// TIA Portal project "Task 1 Faceplate" (V16)

(* hardware
DEVICE "S7-1200 station_1"  S7-1200 Station
   slot 0: "Rack_0"  S7-1200 Rack  Rack  V1.0
   slot 1: "PLC_1"  CPU 1215C DC/DC/DC  6ES7 215-1AG40-0XB0  V4.4
DEVICE "HMI_1"  TP700 Comfort
   slot 0: "HMI_1"  TP700 Comfort  6AV2 124-0GC01-0AX0  16.0.0.0
   slot 1: "HMI_RT_1"  TP700 Comfort  6AV2 124-0GC01-0AX0  16.0.0.0
   slot 5: "HMI_1.IE_CP_1"  PROFINET Interface  16.0.0.0
      slot 1: "PROFINET Interface_1"  PROFINET Interface
         slot 1: "Port_1"  Port
         slot 2: "Port_2"  Port
   slot 7: "HMI_1.MPI/DP_CP_1"  MPI/DP Interface  16.0.0.0
*)

// ===== PLC "PLC_1"  CPU 1215C DC/DC/DC =====

DATA_BLOCK "TASK2 FB"   // DB1
{ S7_Optimized_Access := 'TRUE' }
VERSION : 0.1
// stored: InstanceOfName TASK2
"TASK2"
BEGIN
END_DATA_BLOCK

DATA_BLOCK "TASK1 FB"   // DB2
{ S7_Optimized_Access := 'TRUE' }
VERSION : 0.1
// stored: InstanceOfName TASK1
"TASK1"
BEGIN
END_DATA_BLOCK

DATA_BLOCK "TASK1 DB"   // DB3
{ S7_Optimized_Access := 'TRUE' }
VERSION : 0.1
   VAR
      start : Bool;
      stop : Bool;
      heater : Bool;
   END_VAR
   VAR RETAIN
      temperature : Real;
   END_VAR
   VAR
      run : Bool;
      "max temp" : Real := 50.0;
      "min temp" : Real := 0.0;
      "reset temp" : Real := 0.0;
      reset : Bool;
   END_VAR
   VAR RETAIN
      "preset timer" : DInt := 1000;
   END_VAR
   VAR
      "max limit" : Bool;
      "min limit" : Bool;
      timer_1 : IEC_TIMER;
   END_VAR
BEGIN
END_DATA_BLOCK

DATA_BLOCK "TASK2 DB"   // DB4
{ S7_Optimized_Access := 'TRUE' }
VERSION : 0.1
   VAR
      START : Bool;
      STOP : Bool;
      RUN : Bool;
      FVV : Real := 0.0;
      DVV : Real := 0.0;
      "TIMER" : IEC_TIMER;
      "PRESET TIMER" : Real;
      "MULTIPLY BY X" : Real;
      "MAX LIQUID" : Real := 100.0;
      "MIN LIQUID" : Real := 0.0;
      "H LIQUID ALARM" : Real := 100.0;
      "L LIQUID ALARM" : Real := 20.0;
   END_VAR
BEGIN
END_DATA_BLOCK

FUNCTION_BLOCK "TASK1"   // FB1, LAD
{ S7_Optimized_Access := 'TRUE' }
VERSION : 0.1
   VAR_INPUT
      Start : Bool;
      Stop : Bool;
      reset : Bool;
      "Timer" : DInt;   // value in milliseconds
      "max temperature" : Real;   // max temperature you want in the tank
      "min temperature" : Real;   // min temperature you want in the tank
      "reset temp" : Real;   // to reset the temperature
      "any value" : Real;
      manual : Bool;
   END_VAR
   VAR_OUTPUT
      Output_1 : Bool;
   END_VAR
   VAR_IN_OUT
      Run : Bool;   // process is working
      Heater : Bool;
      "max limit" : Bool;
      "min limit" : Bool;
      Temperature : Real;
      IEC_Timer_0_Instance : TON_TIME;
   END_VAR
   VAR
      Ton : Bool;
      Toff : Bool;   // reset the timer
   END_VAR
BEGIN

REGION Network 1: control operarion
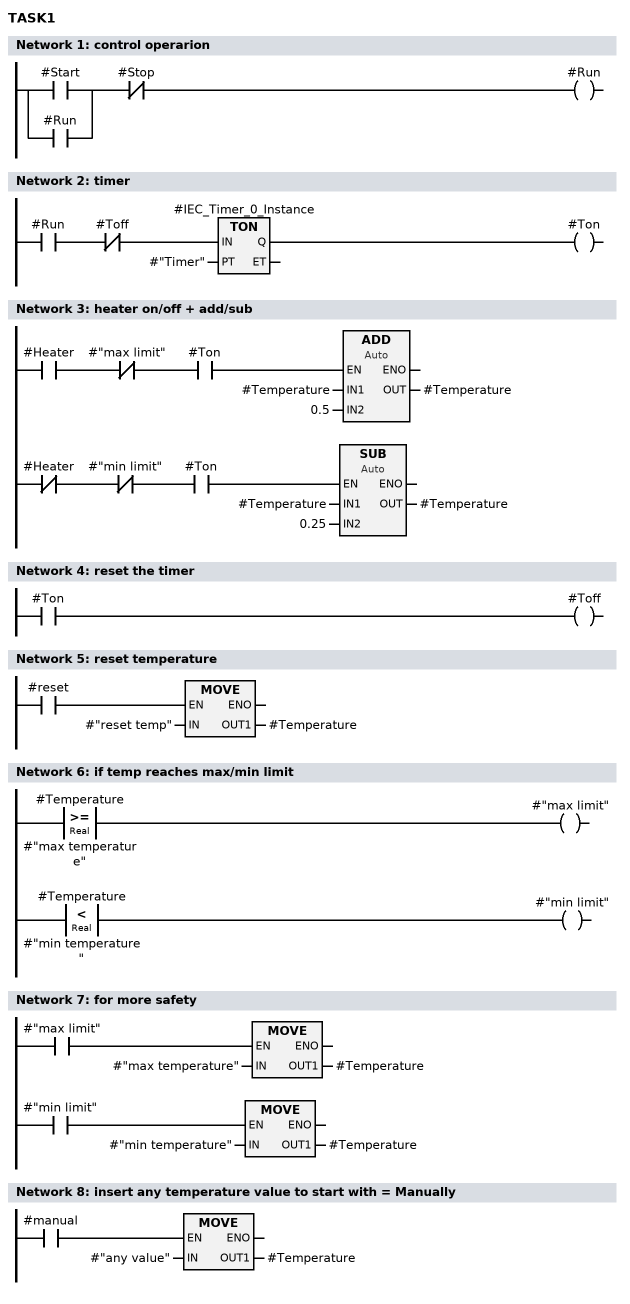
   RUNG wire#powerrail
      Contact( #Start )
      wire#w1
      I_Contact( #Stop )
      Coil( #Run )
   END_RUNG
   RUNG wire#powerrail
      Contact( #Run )
   END_RUNG wire#w1
   // the same network as SCL:
   #Run := (#Start OR #Run) AND NOT #Stop;
END_REGION

REGION Network 2: timer
   #IEC_Timer_0_Instance(IN := #Run AND NOT #Toff, PT := #"Timer");   // TON
   #Ton := #IEC_Timer_0_Instance.Q;
END_REGION

REGION Network 3: heater on/off + add/sub
   RUNG wire#powerrail
      Contact( #Heater )
      I_Contact( #"max limit" )
      Contact( #Ton )
      Add(in1 := #Temperature, in2 := 0.5, out => #Temperature)
   END_RUNG
   RUNG wire#powerrail
      I_Contact( #Heater )
      I_Contact( #"min limit" )
      Contact( #Ton )
      Sub(in1 := #Temperature, in2 := 0.25, out => #Temperature)
   END_RUNG
   // the same network as SCL:
   IF #Heater AND NOT #"max limit" AND #Ton THEN #Temperature := #Temperature + 0.5; END_IF;
   IF NOT #Heater AND NOT #"min limit" AND #Ton THEN #Temperature := #Temperature - 0.25; END_IF;
END_REGION

REGION Network 4: reset the timer
   RUNG wire#powerrail
      Contact( #Ton )
      Coil( #Toff )
   END_RUNG
   // the same network as SCL:
   #Toff := #Ton;
END_REGION

REGION Network 5: reset temperature
   RUNG wire#powerrail
      Contact( #reset )
      Move(in := #"reset temp", out1 => #Temperature)
   END_RUNG
   // the same network as SCL:
   IF #reset THEN #Temperature := #"reset temp"; END_IF;
END_REGION

REGION Network 6: if temp reaches max/min limit
   RUNG wire#powerrail
      { S7_Templates := "SrcType := Real" } GE_Contact(in1 := #Temperature, in2 := #"max temperature")
      Coil( #"max limit" )
   END_RUNG
   RUNG wire#powerrail
      { S7_Templates := "SrcType := Real" } LT_Contact(in1 := #Temperature, in2 := #"min temperature")
      Coil( #"min limit" )
   END_RUNG
   // the same network as SCL:
   #"max limit" := #Temperature >= #"max temperature";
   #"min limit" := #Temperature < #"min temperature";
END_REGION

REGION Network 7: for more safety
   RUNG wire#powerrail
      Contact( #"max limit" )
      Move(in := #"max temperature", out1 => #Temperature)
   END_RUNG
   RUNG wire#powerrail
      Contact( #"min limit" )
      Move(in := #"min temperature", out1 => #Temperature)
   END_RUNG
   // the same network as SCL:
   IF #"max limit" THEN #Temperature := #"max temperature"; END_IF;
   IF #"min limit" THEN #Temperature := #"min temperature"; END_IF;
END_REGION

REGION Network 8: insert any temperature value to start with = Manually
   RUNG wire#powerrail
      Contact( #manual )
      Move(in := #"any value", out1 => #Temperature)
   END_RUNG
   // the same network as SCL:
   IF #manual THEN #Temperature := #"any value"; END_IF;
END_REGION
END_FUNCTION_BLOCK

FUNCTION_BLOCK "TASK2"   // FB2, LAD
{ S7_Optimized_Access := 'TRUE' }
VERSION : 0.1
   VAR_INPUT
      start : Bool;
      stop : Bool;
      "fill valve voltage" : Real;   // analog input from 0-10v
      "drain valve voltage" : Real;   // analog input from 0-10v
      "multiply by x" : Real;   // your max value
      "TIMER" : DInt;   // TIME IN MILLISECONDS FOR CHANGE
      "HIGH LIQUID ALARM" : Real;
      "LOW LIQUID ALARM" : Real;
   END_VAR
   VAR_OUTPUT
      "REAL FVV" : Real;   // real fill valve voltage
      "REAL DVV" : Real;   // real drain valve voltage
      "HIGH LEVEL ALARM" : Bool;
      "LOW LEVEL ALARM" : Bool;
   END_VAR
   VAR_IN_OUT
      run : Bool;
      Rate : Real;   // FLOW OF LIQUID PER TIME
      "REAL FVV - REAL DVV" : Real;
      IEC_Timer_0_Instance : TON_TIME;
      "MAX LEVEL" : Bool;
      "MIN LEVEL" : Bool;
      LEVEL : Real;   // LEVEL OF THE LIQUID
      "MAX LIQUID" : Real;   // MAX LEVEL LIQUID ACCEPTED
      "MIN LIQUID" : Real;   // MIN LEVEL LIQUID ACCEPTED
   END_VAR
   VAR
      "division by 10" : Real := 10.0;
      "FVV after division" : Real;
      "DVV after division" : Real;
      TON : Bool;
      TOFF : Bool;
   END_VAR
BEGIN

REGION Network 1: control process
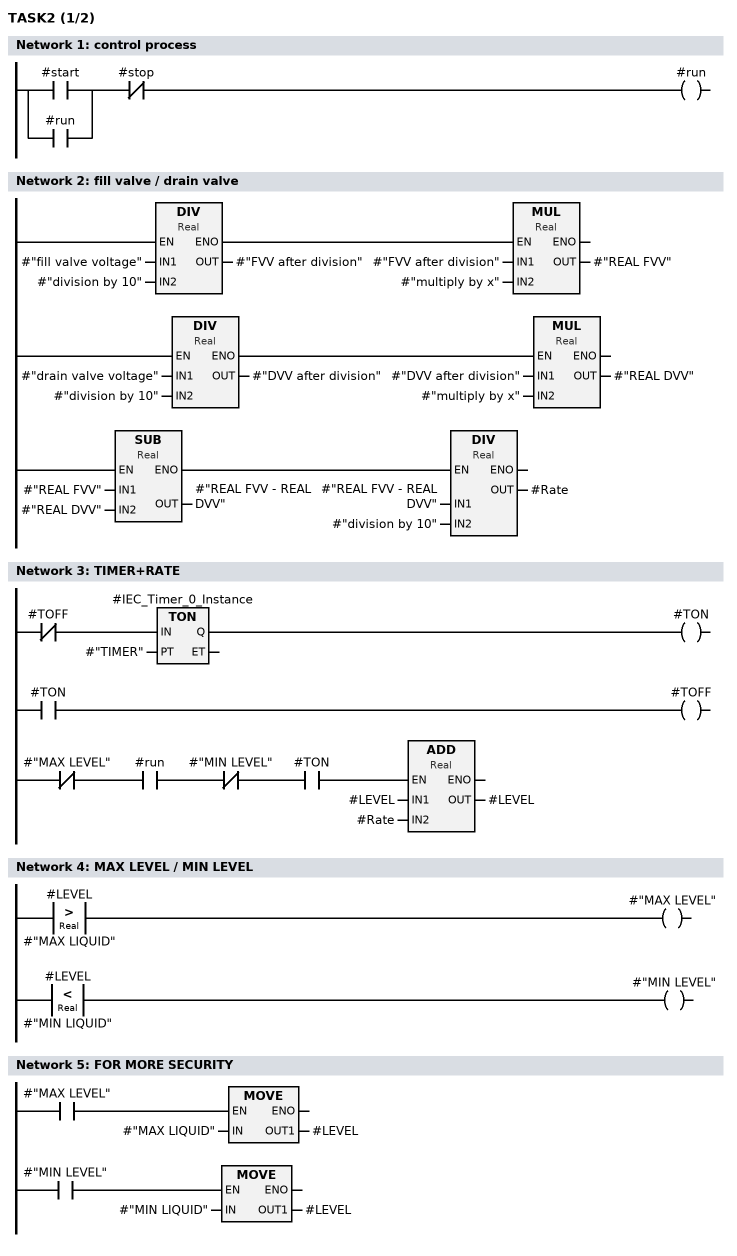
   RUNG wire#powerrail
      Contact( #start )
      wire#w1
      I_Contact( #stop )
      Coil( #run )
   END_RUNG
   RUNG wire#powerrail
      Contact( #run )
   END_RUNG wire#w1
   // the same network as SCL:
   #run := (#start OR #run) AND NOT #stop;
END_REGION

REGION Network 2: fill valve / drain valve
   RUNG wire#powerrail
      { S7_Templates := "SrcType := Real" } Div(in1 := #"fill valve voltage", in2 := #"division by 10", out => #"FVV after division")
      { S7_Templates := "SrcType := Real" } Mul(in1 := #"FVV after division", in2 := #"multiply by x", out => #"REAL FVV")
   END_RUNG
   RUNG wire#powerrail
      { S7_Templates := "SrcType := Real" } Div(in1 := #"drain valve voltage", in2 := #"division by 10", out => #"DVV after division")
      { S7_Templates := "SrcType := Real" } Mul(in1 := #"DVV after division", in2 := #"multiply by x", out => #"REAL DVV")
   END_RUNG
   RUNG wire#powerrail
      { S7_Templates := "SrcType := Real" } Sub(in1 := #"REAL FVV", in2 := #"REAL DVV", out => #"REAL FVV - REAL DVV")
      { S7_Templates := "SrcType := Real" } Div(in1 := #"REAL FVV - REAL DVV", in2 := #"division by 10", out => #Rate)
   END_RUNG
   // the same network as SCL:
   #"FVV after division" := #"fill valve voltage" / #"division by 10";
   #"REAL FVV" := #"FVV after division" * #"multiply by x";
   #"DVV after division" := #"drain valve voltage" / #"division by 10";
   #"REAL DVV" := #"DVV after division" * #"multiply by x";
   #"REAL FVV - REAL DVV" := #"REAL FVV" - #"REAL DVV";
   #Rate := #"REAL FVV - REAL DVV" / #"division by 10";
END_REGION

REGION Network 3: TIMER+RATE
   #IEC_Timer_0_Instance(IN := NOT #TOFF, PT := #"TIMER");   // TON
   #TON := #IEC_Timer_0_Instance.Q;
   #TOFF := #TON;
   IF NOT #"MAX LEVEL" AND #run AND NOT #"MIN LEVEL" AND #TON THEN #LEVEL := #LEVEL + #Rate; END_IF;
END_REGION

REGION Network 4: MAX LEVEL / MIN LEVEL
   RUNG wire#powerrail
      { S7_Templates := "SrcType := Real" } GT_Contact(in1 := #LEVEL, in2 := #"MAX LIQUID")
      Coil( #"MAX LEVEL" )
   END_RUNG
   RUNG wire#powerrail
      { S7_Templates := "SrcType := Real" } LT_Contact(in1 := #LEVEL, in2 := #"MIN LIQUID")
      Coil( #"MIN LEVEL" )
   END_RUNG
   // the same network as SCL:
   #"MAX LEVEL" := #LEVEL > #"MAX LIQUID";
   #"MIN LEVEL" := #LEVEL < #"MIN LIQUID";
END_REGION

REGION Network 5: FOR MORE SECURITY
   RUNG wire#powerrail
      Contact( #"MAX LEVEL" )
      Move(in := #"MAX LIQUID", out1 => #LEVEL)
   END_RUNG
   RUNG wire#powerrail
      Contact( #"MIN LEVEL" )
      Move(in := #"MIN LIQUID", out1 => #LEVEL)
   END_RUNG
   // the same network as SCL:
   IF #"MAX LEVEL" THEN #LEVEL := #"MAX LIQUID"; END_IF;
   IF #"MIN LEVEL" THEN #LEVEL := #"MIN LIQUID"; END_IF;
END_REGION

REGION Network 6: HIGH LEVEL ALARM / LOW LEVEL ALARM
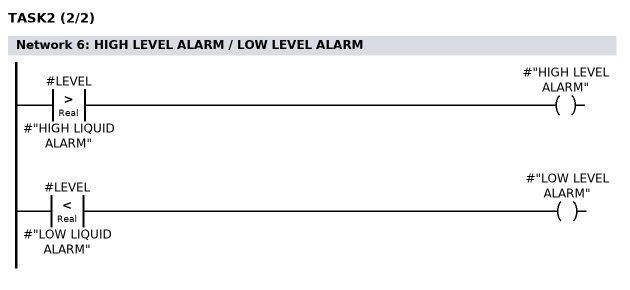
   RUNG wire#powerrail
      { S7_Templates := "SrcType := Real" } GT_Contact(in1 := #LEVEL, in2 := #"HIGH LIQUID ALARM")
      Coil( #"HIGH LEVEL ALARM" )
   END_RUNG
   RUNG wire#powerrail
      { S7_Templates := "SrcType := Real" } LT_Contact(in1 := #LEVEL, in2 := #"LOW LIQUID ALARM")
      Coil( #"LOW LEVEL ALARM" )
   END_RUNG
   // the same network as SCL:
   #"HIGH LEVEL ALARM" := #LEVEL > #"HIGH LIQUID ALARM";
   #"LOW LEVEL ALARM" := #LEVEL < #"LOW LIQUID ALARM";
END_REGION
END_FUNCTION_BLOCK

ORGANIZATION_BLOCK "Main"   // OB1, LAD, ProgramCycle
TITLE = "Main Program Sweep (Cycle)"
{ S7_Optimized_Access := 'TRUE' }
VERSION : 0.1
   VAR_INPUT
      Initial_Call : Bool;   // Initial call of this OB
      Remanence : Bool;   // =True, if remanent data are available
   END_VAR
BEGIN

REGION Network 1
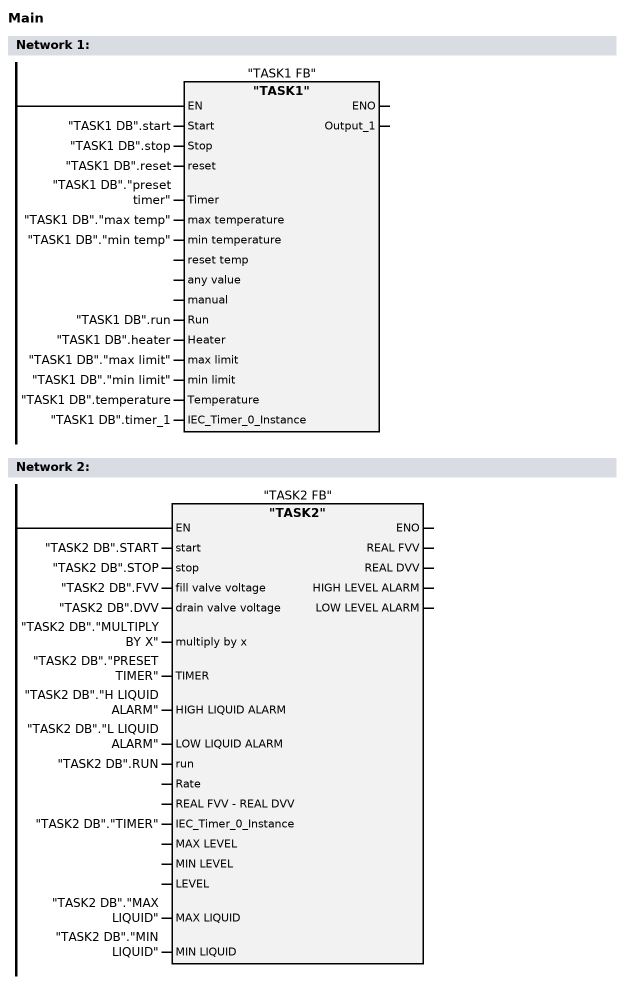
   RUNG wire#powerrail
      "TASK1 FB"(Start := "TASK1 DB".start, Stop := "TASK1 DB".stop, reset := "TASK1 DB".reset, "Timer" := "TASK1 DB"."preset timer", "max temperature" := "TASK1 DB"."max temp", "min temperature" := "TASK1 DB"."min temp", "reset temp" :=, "any value" :=, manual :=, Run := "TASK1 DB".run, Heater := "TASK1 DB".heater, "max limit" := "TASK1 DB"."max limit", "min limit" := "TASK1 DB"."min limit", Temperature := "TASK1 DB".temperature, IEC_Timer_0_Instance := "TASK1 DB".timer_1, Output_1 =>)
   END_RUNG
   // the same network as SCL:
   "TASK1 FB"(Start := "TASK1 DB".start,   // "TASK1"
              Stop := "TASK1 DB".stop,
              reset := "TASK1 DB".reset,
              "Timer" := "TASK1 DB"."preset timer",
              "max temperature" := "TASK1 DB"."max temp",
              "min temperature" := "TASK1 DB"."min temp",
              Run := "TASK1 DB".run,
              Heater := "TASK1 DB".heater,
              "max limit" := "TASK1 DB"."max limit",
              "min limit" := "TASK1 DB"."min limit",
              Temperature := "TASK1 DB".temperature,
              IEC_Timer_0_Instance := "TASK1 DB".timer_1);
END_REGION

REGION Network 2
   RUNG wire#powerrail
      "TASK2 FB"(start := "TASK2 DB".START, stop := "TASK2 DB".STOP, "fill valve voltage" := "TASK2 DB".FVV, "drain valve voltage" := "TASK2 DB".DVV, "multiply by x" := "TASK2 DB"."MULTIPLY BY X", "TIMER" := "TASK2 DB"."PRESET TIMER", "HIGH LIQUID ALARM" := "TASK2 DB"."H LIQUID ALARM", "LOW LIQUID ALARM" := "TASK2 DB"."L LIQUID ALARM", run := "TASK2 DB".RUN, Rate :=, "REAL FVV - REAL DVV" :=, IEC_Timer_0_Instance := "TASK2 DB"."TIMER", "MAX LEVEL" :=, "MIN LEVEL" :=, LEVEL :=, "MAX LIQUID" := "TASK2 DB"."MAX LIQUID", "MIN LIQUID" := "TASK2 DB"."MIN LIQUID", "REAL FVV" =>, "REAL DVV" =>, "HIGH LEVEL ALARM" =>, "LOW LEVEL ALARM" =>)
   END_RUNG
   // the same network as SCL:
   "TASK2 FB"(start := "TASK2 DB".START,   // "TASK2"
              stop := "TASK2 DB".STOP,
              "fill valve voltage" := "TASK2 DB".FVV,
              "drain valve voltage" := "TASK2 DB".DVV,
              "multiply by x" := "TASK2 DB"."MULTIPLY BY X",
              "TIMER" := "TASK2 DB"."PRESET TIMER",
              "HIGH LIQUID ALARM" := "TASK2 DB"."H LIQUID ALARM",
              "LOW LIQUID ALARM" := "TASK2 DB"."L LIQUID ALARM",
              run := "TASK2 DB".RUN,
              IEC_Timer_0_Instance := "TASK2 DB"."TIMER",
              "MAX LIQUID" := "TASK2 DB"."MAX LIQUID",
              "MIN LIQUID" := "TASK2 DB"."MIN LIQUID");
END_REGION
END_ORGANIZATION_BLOCK

// ===== library: MasterCopy "TASK1 DB" =====

DATA_BLOCK "TASK1 DB"   // DB3
{ S7_Optimized_Access := 'TRUE' }
VERSION : 0.1
   VAR
      start : Bool;
      stop : Bool;
      heater : Bool;
   END_VAR
   VAR RETAIN
      temperature : Real;
   END_VAR
   VAR
      run : Bool;
      "max temp" : Real := 50.0;
      "min temp" : Real := 0.0;
      "reset temp" : Real := 0.0;
      reset : Bool;
   END_VAR
   VAR RETAIN
      "preset timer" : DInt := 1000;
   END_VAR
   VAR
      "max limit" : Bool;
      "min limit" : Bool;
      timer_1 : IEC_TIMER;
   END_VAR
BEGIN
END_DATA_BLOCK

// ===== library: MasterCopy "TASK2 DB" =====

DATA_BLOCK "TASK2 DB"   // DB4
{ S7_Optimized_Access := 'TRUE' }
VERSION : 0.1
   VAR
      START : Bool;
      STOP : Bool;
      RUN : Bool;
      FVV : Real := 0.0;
      DVV : Real := 0.0;
      "TIMER" : IEC_TIMER;
      "PRESET TIMER" : Real;
      "MULTIPLY BY X" : Real;
      "MAX LIQUID" : Real := 100.0;
      "MIN LIQUID" : Real := 0.0;
      "H LIQUID ALARM" : Real := 100.0;
      "L LIQUID ALARM" : Real := 20.0;
   END_VAR
BEGIN
END_DATA_BLOCK

(* ===== HMI "HMI_RT_1" =====
system functions are stored by id; their names below are inferred from use
connection "HMI_Connection_1": ETHERNET, S7_1200_OMS

HMI tags "Default tag table"
   "Tag_ScreenNumber" : UInt, internal
   "Data_block_1_temperature" : Real = PLC "TASK1 DB".temperature, 1 s
   "Data_block_1_start" : Bool = PLC "TASK1 DB".start, 1 s
   "Data_block_1_heater" : Bool = PLC "TASK1 DB".heater, 1 s
   "TASK1 DB_stop" : Bool = PLC "TASK1 DB".stop, 1 s
   "TASK1 DB_reset" : Bool = PLC "TASK1 DB".reset, 1 s

Template "Template_1" 800x480
   Button "Exit" at 714,429 size 71x50; TextOff 'Exit'; PictureOff "ExitRuntime_KTP700_Basic_PN_TR"; PictureOn "ExitRuntime_KTP700_Basic_PN_TR"
      on Release: StopRuntime(0)
   Button "Template_Button" at 614,429 size 71x50; TextOff 'Text'
   Button "Template_Button_1" at 514,429 size 71x50; TextOff 'Text'
   Button "Template_Button_2" at 414,429 size 71x50; TextOff 'Text'
   Button "Template_Button_3" at 314,429 size 71x50; TextOff 'Text'
   Button "Template_Button_4" at 214,429 size 71x50; TextOff 'Text'
   Button "Template_Button_5" at 114,429 size 71x50; TextOff 'Text'
   Button "Start screen" at 14,429 size 71x50; TextOff 'Start screen'; PictureOff "NavigateHome_KTP700_Basic_PN_TR"; PictureOn "NavigateHome_KTP700_Basic_PN_TR"
      on Release: ActivateScreen("Root screen", 0)
   SymbolicIOField "Symbolic_IO_Field_Screen" at 93,9 size 600x33; TextOff '0'; TextOn '1'; TextList "TextList_ScreenNames"
      ProcessValue <- "Tag_ScreenNumber"
      on Change: ActivateScreenByNumber("Tag_ScreenNumber", 0)
   DateTimeField "HmiScreenItemData" at 695,25 size 105x25
   DateTimeField "HmiScreenItemData_1" at 695,0 size 105x25
   GraphicView "Logo" at 0,0 size 91x51; Picture "Logo of HMI_1"

screen "Root screen" 800x480, template "Template_1"
   on GenerateScreen: SetTag("Tag_ScreenNumber", 1)
   TextField "HmiScreenItemData" at 86,12 size 640x25; Text 'Welcome to HMI_1 (KTP700 Basic+ PN)!'
   ScreenModuleView "Faceplate_3_1" at 50,59 size 202x216; Guid_{11997190-8919} 'temp1'; ScreenModuleType ""; Guid_{11997190-9122} 'Temperature'
      Guid_{11997190-7705} <- "Data_block_1_heater"
      Guid_{11997190-7699} <- "Data_block_1_start"
      Guid_{11997190-7703} <- "TASK1 DB_stop"
      Guid_{11997190-7872} <- "Data_block_1_temperature"
      Guid_{11997190-7707} <- "TASK1 DB_reset"
   ScreenModuleView "Faceplate_3_2" at 297,56 size 202x216; ScreenModuleType ""
      Guid_{11997190-7705} <- "Data_block_1_heater"
*)

(* ===== HMI "HMI_RT_1" =====

ScreenModuleEditorView "Faceplate_3" 640x480
   Button "Button_2" at 14,148 size 96x32; TextOff 'Start'
   Button "Button_3" at 115,148 size 96x32; TextOff 'Stop'
   IOField "I/O field_1" at 31,56 size 165x32; FormatPattern s999.99
   Button "Button_4" at 53,17 size 116x32; TextOff 'Temperature'
   Switch "Switch_1" at 51,102 size 114x32; TextOn 'Heater ON'; CaptionText 'Switch'; TextOff 'Heater OFF'
   Button "Button_1" at 59,192 size 96x32; TextOff 'Reset'
*)

(* ===== HMI "HMI_RT_1" =====

ScreenModuleEditorView "Faceplate_3" 640x480
   Button "Button_2" at 14,148 size 96x32; TextOff 'Start'
   Button "Button_3" at 115,148 size 96x32; TextOff 'Stop'
   IOField "I/O field_1" at 31,56 size 165x32; FormatPattern s999.99
   Button "Button_4" at 53,17 size 116x32; TextOff 'Temperature'
   Switch "Switch_1" at 51,102 size 114x32; TextOn 'Heater ON'; CaptionText 'Switch'; TextOff 'Heater OFF'
   Button "Button_1" at 59,192 size 96x32; TextOff 'Reset'
*)

(* ===== HMI "HMI_RT_1" =====

ScreenModuleEditorView "Faceplate_3" 640x480
   Button "Button_2" at 14,148 size 96x32; TextOff 'Start'
   Button "Button_3" at 115,148 size 96x32; TextOff 'Stop'
   IOField "I/O field_1" at 31,56 size 165x32; FormatPattern s999.99
   Button "Button_4" at 53,17 size 116x32; TextOff 'Temperature'
   Switch "Switch_1" at 51,102 size 114x32; TextOn 'Heater ON'; CaptionText 'Switch'; TextOff 'Heater OFF'
   Button "Button_1" at 59,192 size 96x32; TextOff 'Reset'
*)

(* ===== HMI "HMI_RT_1" =====
system functions are stored by id; their names below are inferred from use

ScreenModuleEditorView "Faceplate_3" 640x480
   Button "Button_2" at 14,148 size 96x32; TextOff 'Start'
      on Press: SetBit("Start")
      on Release: ResetBit("Start")
   Button "Button_3" at 115,148 size 96x32; TextOff 'Stop'
      ProcessValue <- "stop"
      on Press: SetBit("stop")
      on Release: ResetBit("stop")
   IOField "I/O field_1" at 31,56 size 165x32; FormatPattern s99999
      ProcessValue <- "Temperature"
   Button "Button_4" at 44,17 size 130x32; TextOff 'Temperature'
   Switch "Switch_1" at 51,102 size 114x32; TextOn 'Heater ON'; CaptionText 'Switch'; TextOff 'Heater OFF'
      on SwitchOn: SetBit("Heater")
      on SwitchOff: ResetBit("Heater")
   Button "Button_1" at 59,192 size 96x32; TextOff 'Reset'
*)

(* ===== HMI "HMI_RT_1" =====
system functions are stored by id; their names below are inferred from use

ScreenModuleEditorView "Faceplate_3" 640x480
   Button "Button_2" at 14,148 size 96x32; TextOff 'Start'
      on Release: ResetBit("Start")
      on Press: SetBit("Start")
   Button "Button_3" at 115,148 size 96x32; TextOff 'Stop'
      on Release: ResetBit("stop")
      on Press: SetBit("stop")
      ProcessValue <- "stop"
   IOField "I/O field_1" at 31,56 size 165x32; FormatPattern s99999
      ProcessValue <- "Temperature"
   Button "Button_4" at 44,17 size 130x32; TextOff 'Temperature'
   Switch "Switch_1" at 51,102 size 114x32; TextOn 'Heater ON'; CaptionText 'Switch'; TextOff 'Heater OFF'
      on SwitchOff: ResetBit("Heater")
      on SwitchOn: SetBit("Heater")
   Button "Button_1" at 59,192 size 96x32; TextOff 'Reset'
*)

(* ===== HMI "HMI_RT_1" =====
system functions are stored by id; their names below are inferred from use

ScreenModuleEditorView "Faceplate_3" 640x480
   Button "Button_2" at 14,148 size 96x32; TextOff 'Start'
      on Release: ResetBit("Start")
      on Press: SetBit("Start")
      ProcessValue <- "Start"
   Button "Button_3" at 115,148 size 96x32; TextOff 'Stop'
      on Release: ResetBit("stop")
      on Press: SetBit("stop")
      ProcessValue <- "stop"
   IOField "I/O field_1" at 31,56 size 165x32; FormatPattern s99999
      ProcessValue <- "Temperature"
   Button "Button_4" at 44,17 size 130x32; TextOff 'Temperature'
   Switch "Switch_1" at 51,102 size 114x32; TextOn 'Heater ON'; CaptionText 'Switch'; TextOff 'Heater OFF'
      on SwitchOn: SetBit("Heater")
      on SwitchOff: ResetBit("Heater")
      ProcessValue <- "Heater"
   Button "Button_1" at 59,192 size 96x32; TextOff 'Reset'
      ProcessValue <- "reset"
*)

(* ===== HMI "HMI_RT_1" =====
system functions are stored by id; their names below are inferred from use

ScreenModuleEditorView "Faceplate_3" 640x480
   Button "Button_2" at 14,148 size 96x32; TextOff 'Start'
      on Release: ResetBit("Start")
      on Press: SetBit("Start")
      ProcessValue <- "Start"
   Button "Button_3" at 115,148 size 96x32; TextOff 'Stop'
      on Release: ResetBit("stop")
      on Press: SetBit("stop")
      ProcessValue <- "stop"
   IOField "I/O field_1" at 31,56 size 165x32; FormatPattern s999.99
      ProcessValue <- "Temperature"
   Button "Button_4" at 44,17 size 130x32; TextOff 'Temperature'
   Switch "Switch_1" at 51,102 size 114x32; TextOn 'Heater ON'; CaptionText 'Switch'; TextOff 'Heater OFF'
      on SwitchOff: ResetBit("Heater")
      on SwitchOn: SetBit("Heater")
      ProcessValue <- "Heater"
   Button "Button_1" at 59,192 size 96x32; TextOff 'Reset'
      ProcessValue <- "reset"
*)

(* ===== HMI "HMI_RT_1" =====
system functions are stored by id; their names below are inferred from use

ScreenModuleEditorView "Faceplate_3" 640x480
   Button "Button_2" at 14,148 size 96x32; TextOff 'Start'
      on Release: ResetBit("Start")
      on Press: SetBit("Start")
      ProcessValue <- "Start"
   Button "Button_3" at 115,148 size 96x32; TextOff 'Stop'
      on Release: ResetBit("stop")
      on Press: SetBit("stop")
      ProcessValue <- "stop"
   IOField "I/O field_1" at 31,56 size 165x32; FormatPattern s999.99
      ProcessValue <- "Temperature"
   Button "Button_4" at 44,17 size 130x32; TextOff 'Temperature'
   Switch "Switch_1" at 51,102 size 114x32; TextOn 'Heater ON'; CaptionText 'Switch'; TextOff 'Heater OFF'
      on SwitchOff: ResetBit("Heater")
      on SwitchOn: SetBit("Heater")
      ProcessValue <- "Heater"
   Button "Button_1" at 59,192 size 96x32; TextOff 'Reset'
      ProcessValue <- "reset"
      on Press: SetBit("reset")
      on Release: ResetBit("reset")
*)

(* ===== HMI "HMI_RT_1" =====
system functions are stored by id; their names below are inferred from use

ScreenModuleEditorView "Faceplate_3" 640x480
   Button "Button_2" at 14,148 size 96x32; TextOff 'Start'
      on Release: ResetBit("Start")
      on Press: SetBit("Start")
      ProcessValue <- "Start"
   Button "Button_3" at 115,148 size 96x32; TextOff 'Stop'
      on Release: ResetBit("stop")
      on Press: SetBit("stop")
      ProcessValue <- "stop"
   IOField "I/O field_1" at 31,56 size 165x32; FormatPattern s999.99
      ProcessValue <- "Temperature"
   Button "Button_4" at 44,17 size 130x32; TextOff 'Temperature'
   Switch "Switch_1" at 51,102 size 114x32; TextOn 'Heater ON'; CaptionText 'Switch'; TextOff 'Heater OFF'
      on SwitchOff: ResetBit("Heater")
      on SwitchOn: SetBit("Heater")
      ProcessValue <- "Heater"
      Appearance <- "Heater"
   Button "Button_1" at 59,192 size 96x32; TextOff 'Reset'
      on Release: ResetBit("reset")
      on Press: SetBit("reset")
      ProcessValue <- "reset"
*)

(* ===== HMI "HMI_RT_1" =====
system functions are stored by id; their names below are inferred from use

ScreenModuleEditorView "Faceplate_3" 640x480
   Button "Button_2" at 14,148 size 96x32; TextOff 'Start'
      on Release: ResetBit("Start")
      on Press: SetBit("Start")
      ProcessValue <- "Start"
   Button "Button_3" at 115,148 size 96x32; TextOff 'Stop'
      on Release: ResetBit("stop")
      on Press: SetBit("stop")
      ProcessValue <- "stop"
   IOField "I/O field_1" at 31,56 size 165x32; FormatPattern s999.99
      ProcessValue <- "Temperature"
   Button "Button_4" at 44,17 size 130x32; TextOff 'Temperature'
   Switch "Switch_1" at 51,102 size 114x32; TextOn 'Heater ON'; CaptionText 'Switch'; TextOff 'Heater OFF'
      on SwitchOff: ResetBit("Heater")
      on SwitchOn: SetBit("Heater")
      Appearance <- "Heater"
      ProcessValue <- "Heater"
   Button "Button_1" at 59,192 size 96x32; TextOff 'Reset'
      on Release: ResetBit("reset")
      on Press: SetBit("reset")
      ProcessValue <- "reset"
*)

(* ===== HMI "HMI_RT_1" =====
system functions are stored by id; their names below are inferred from use

ScreenModuleEditorView "Faceplate_3" 640x480
   Button "Button_2" at 14,148 size 96x32; TextOff 'Start'
      on Release: ResetBit("Start")
      on Press: SetBit("Start")
      ProcessValue <- "Start"
   Button "Button_3" at 115,148 size 96x32; TextOff 'Stop'
      on Release: ResetBit("stop")
      on Press: SetBit("stop")
      ProcessValue <- "stop"
   IOField "I/O field_1" at 31,56 size 165x32; FormatPattern s999.99
      ProcessValue <- "Temperature"
   Switch "Switch_1" at 59,104 size 114x32; TextOn 'Heater ON'; CaptionText 'Switch'; TextOff 'Heater OFF'
      on SwitchOff: ResetBit("Heater")
      on SwitchOn: SetBit("Heater")
      Appearance <- "Heater"
      ProcessValue <- "Heater"
   Button "Button_1" at 59,192 size 96x32; TextOff 'Reset'
      on Release: ResetBit("reset")
      on Press: SetBit("reset")
      ProcessValue <- "reset"
   TextField "Text field_1" at 64,24 size 101x22; Text 'Temperature'
*)

(* ===== HMI "HMI_RT_1" =====
system functions are stored by id; their names below are inferred from use

ScreenModuleEditorView "Faceplate_3" 640x480
   Button "Button_2" at 19,101 size 96x32; TextOff 'Start'
      on Release: ResetBit("Start")
      on Press: SetBit("Start")
      ProcessValue <- "Start"
   Button "Button_3" at 116,101 size 96x32; TextOff 'Stop'
      on Release: ResetBit("stop")
      on Press: SetBit("stop")
      ProcessValue <- "stop"
   IOField "I/O field_1" at 31,56 size 165x32; FormatPattern s999.99
      ProcessValue <- "Temperature"
   Switch "Switch_1" at 64,186 size 114x32; TextOn 'Heater ON'; CaptionText 'Switch'; TextOff 'Heater OFF'
      on SwitchOff: ResetBit("Heater")
      on SwitchOn: SetBit("Heater")
      Appearance <- "Heater"
      ProcessValue <- "Heater"
   Button "Button_1" at 68,145 size 96x32; TextOff 'Reset'
      on Release: ResetBit("reset")
      on Press: SetBit("reset")
      ProcessValue <- "reset"
   TextField "Text field_1" at 64,24 size 101x22; Text 'Temperature'
*)